REGION Network 107: DB34.DBB10 -> DB86.DBB20 / 8 y 8
   // Falla Compresor ABC2 Baja Presion de Agua
   // Falla Compresor ABC2 Alta Temperatura de Aire
   // Falla Compresor ABC2 Alta Temperatura de agua
   // Falla Compresor ABC3 Baja Presion de Aceite
   // Falla Compresor ABC3 Baja Presion de Agua
   // Falla Compresor ABC3 Alta Temperatura de Aire
   // Falla Compresor ABC3 Alta Temperatura de agua
   // Falla Compresor ABC4 Baja Presion de Aceite
   RUNG wire#powerrail
      { S7_GenerateENO := "TRUE" } Move(in := %DB34.DBB10, out1 => %DB86.DBB20)
      "And-Byte MTA"(IN0 := %DB86.DBB21, IN1 := %DB34.DBB10, OUT2 => %DB86.DBB21)
      { S7_GenerateENO := "TRUE" } Move(in := %DB86.DBB21, out1 => %DB35.DBB10)
   END_RUNG
   // the same network as SCL:
   // ENO of a box is taken as its EN; it also drops when the box reports an error
   %DB86.DBB20 := %DB34.DBB10;
   "And-Byte MTA"(IN0 := %DB86.DBB21, IN1 := %DB34.DBB10, OUT2 => %DB86.DBB21, ENO => #_w1);
   IF #_w1 THEN %DB35.DBB10 := %DB86.DBB21; END_IF;
END_REGION

REGION Network 108: DB34.DBB11 -> DB86.DBB22 / 8 y 8
   // Falla Compresor ABC4 Alta Temperatura de Aire
   // Falla Compresor ABC4 Alta Temperatura de Aire
   // Falla Compresor ABC4 Alta Temperatura de agua
   // Falla Compresor ABC5 Baja Presion de Aceite
   // Falla Compresor ABC5 Alta Temperatura de Aire
   // Falla Compresor ABC5 Alta Temperatura de Aire
   // Falla Compresor ABC5 Alta Temperatura de agua
   // Falla Compresor Bellis & MHW28 Baja Presion Aceite
   RUNG wire#powerrail
      { S7_GenerateENO := "TRUE" } Move(in := %DB34.DBB11, out1 => %DB86.DBB22)
      "And-Byte MTA"(IN0 := %DB86.DBB23, IN1 := %DB34.DBB11, OUT2 => %DB86.DBB23)
      { S7_GenerateENO := "TRUE" } Move(in := %DB86.DBB23, out1 => %DB35.DBB11)
   END_RUNG
   // the same network as SCL:
   // ENO of a box is taken as its EN; it also drops when the box reports an error
   %DB86.DBB22 := %DB34.DBB11;
   "And-Byte MTA"(IN0 := %DB86.DBB23, IN1 := %DB34.DBB11, OUT2 => %DB86.DBB23, ENO => #_w1);
   IF #_w1 THEN %DB35.DBB11 := %DB86.DBB23; END_IF;
END_REGION

REGION Network 109: DB34.DBB12 -> DB86.DBB24 / 8 y 8
   // Falla Compresor Bellis & MHW28 Baja Presion de Agua
   // Falla Compresor Bellis & MHW28 Alta temperatura de Aire
   // Falla Compresor Bellis & MHW28 Alta temperatura de Agua
   // Falla Compresor Bellis & MHW28 Falla de Flujostato
   // Requiere Marcha MC001
   // Requiere Marcha MC002
   // Requiere Marcha MC003
   // Requiere Marcha MC004
   RUNG wire#powerrail
      { S7_GenerateENO := "TRUE" } Move(in := %DB34.DBB12, out1 => %DB86.DBB24)
      "And-Byte MTA"(IN0 := %DB86.DBB25, IN1 := %DB34.DBB12, OUT2 => %DB86.DBB25)
      { S7_GenerateENO := "TRUE" } Move(in := %DB86.DBB25, out1 => %DB35.DBB12)
   END_RUNG
   // the same network as SCL:
   // ENO of a box is taken as its EN; it also drops when the box reports an error
   %DB86.DBB24 := %DB34.DBB12;
   "And-Byte MTA"(IN0 := %DB86.DBB25, IN1 := %DB34.DBB12, OUT2 => %DB86.DBB25, ENO => #_w1);
   IF #_w1 THEN %DB35.DBB12 := %DB86.DBB25; END_IF;
END_REGION

REGION Network 110: DB34.DBB13 -> DB86.DBB26 / 8 y 8
   // Requiere Marcha MC005
   // Falla Conexión con sensor de Temperatura torres de Cavaleto
   // Falla Conexión con sensor de Temperatura torres de Chillers
   // Falla Conexión con sensor de Presión de ALTA
   // Falla Conexión con sensor de Presión de ALTA redundante
   // Falla Conexión con sensor de Presión de Baja
   // Falla Presión de Alta en Límite Mínimo
   // Falla Presión de Alta en demasiado Baja
   RUNG wire#powerrail
      { S7_GenerateENO := "TRUE" } Move(in := %DB34.DBB13, out1 => %DB86.DBB26)
      "And-Byte MTA"(IN0 := %DB86.DBB27, IN1 := %DB34.DBB13, OUT2 => %DB86.DBB27)
      { S7_GenerateENO := "TRUE" } Move(in := %DB86.DBB27, out1 => %DB35.DBB13)
   END_RUNG
   // the same network as SCL:
   // ENO of a box is taken as its EN; it also drops when the box reports an error
   %DB86.DBB26 := %DB34.DBB13;
   "And-Byte MTA"(IN0 := %DB86.DBB27, IN1 := %DB34.DBB13, OUT2 => %DB86.DBB27, ENO => #_w1);
   IF #_w1 THEN %DB35.DBB13 := %DB86.DBB27; END_IF;
END_REGION

REGION Network 111: DB34.DBB14 -> DB86.DBB28 / 8 y 8
   // Falla Presión de Alta en demasiado Alta
   // Falla Presión de Alta en Límite Máximo
   // Falla Presión de Baja en Límite Mínimo
   // Falla Presión de Baja en demasiado Baja
   // Falla Presión de Baja en demasiado Alta
   // Falla Presión de Baja en Límite Máximo
   // Falla en chiller de envasado chico
   // Falla en chiller de soplado chico
   RUNG wire#powerrail
      { S7_GenerateENO := "TRUE" } Move(in := %DB34.DBB14, out1 => %DB86.DBB28)
      "And-Byte MTA"(IN0 := %DB86.DBB29, IN1 := %DB34.DBB14, OUT2 => %DB86.DBB29)
      { S7_GenerateENO := "TRUE" } Move(in := %DB86.DBB29, out1 => %DB35.DBB14)
   END_RUNG
   // the same network as SCL:
   // ENO of a box is taken as its EN; it also drops when the box reports an error
   %DB86.DBB28 := %DB34.DBB14;
   "And-Byte MTA"(IN0 := %DB86.DBB29, IN1 := %DB34.DBB14, OUT2 => %DB86.DBB29, ENO => #_w1);
   IF #_w1 THEN %DB35.DBB14 := %DB86.DBB29; END_IF;
END_REGION

REGION Network 112: DB34.DBB15 -> DB86.DBB30 / 8 y 8
   // Horas máximas en Compresor 1
   // Horas máximas en Compresor 2
   // Horas máximas en Compresor 3
   // Horas máximas en Compresor 4
   // Horas máximas en Compresor 5
   // Falla algún contactor en Booster 1
   // Falla algún guardamotor en Booster 1
   // Presión Alta en Booster
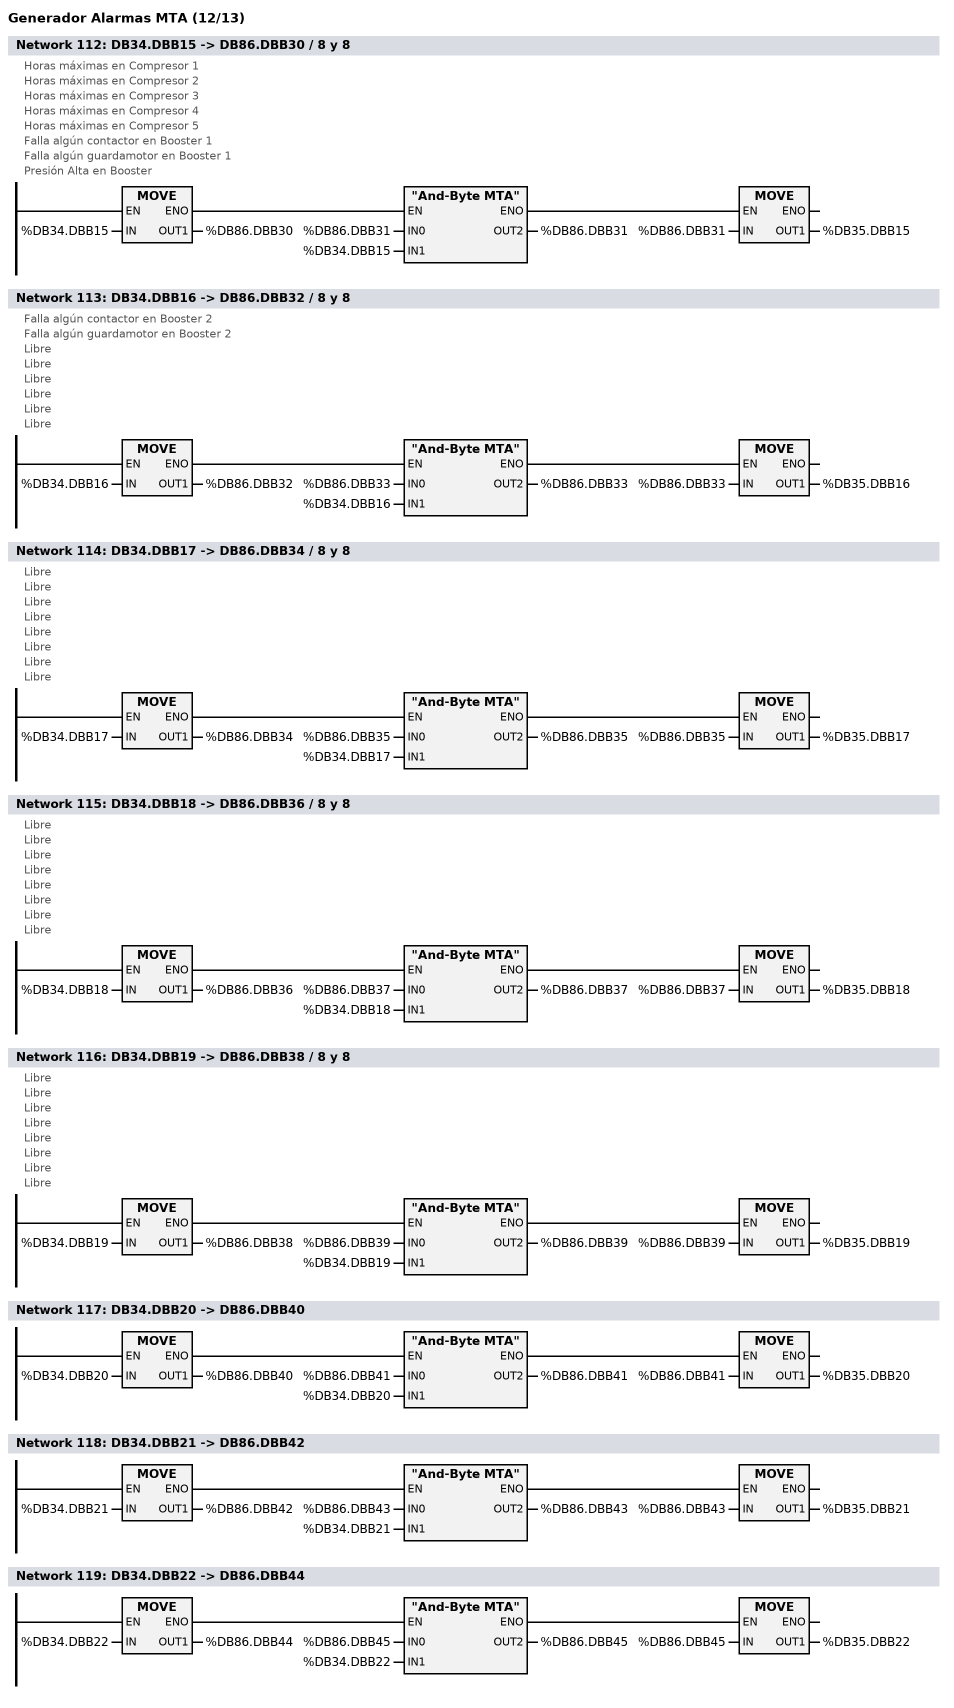
   RUNG wire#powerrail
      { S7_GenerateENO := "TRUE" } Move(in := %DB34.DBB15, out1 => %DB86.DBB30)
      "And-Byte MTA"(IN0 := %DB86.DBB31, IN1 := %DB34.DBB15, OUT2 => %DB86.DBB31)
      { S7_GenerateENO := "TRUE" } Move(in := %DB86.DBB31, out1 => %DB35.DBB15)
   END_RUNG
   // the same network as SCL:
   // ENO of a box is taken as its EN; it also drops when the box reports an error
   %DB86.DBB30 := %DB34.DBB15;
   "And-Byte MTA"(IN0 := %DB86.DBB31, IN1 := %DB34.DBB15, OUT2 => %DB86.DBB31, ENO => #_w1);
   IF #_w1 THEN %DB35.DBB15 := %DB86.DBB31; END_IF;
END_REGION

REGION Network 113: DB34.DBB16 -> DB86.DBB32 / 8 y 8
   // Falla algún contactor en Booster 2
   // Falla algún guardamotor en Booster 2
   // Libre
   // Libre
   // Libre
   // Libre
   // Libre
   // Libre
   RUNG wire#powerrail
      { S7_GenerateENO := "TRUE" } Move(in := %DB34.DBB16, out1 => %DB86.DBB32)
      "And-Byte MTA"(IN0 := %DB86.DBB33, IN1 := %DB34.DBB16, OUT2 => %DB86.DBB33)
      { S7_GenerateENO := "TRUE" } Move(in := %DB86.DBB33, out1 => %DB35.DBB16)
   END_RUNG
   // the same network as SCL:
   // ENO of a box is taken as its EN; it also drops when the box reports an error
   %DB86.DBB32 := %DB34.DBB16;
   "And-Byte MTA"(IN0 := %DB86.DBB33, IN1 := %DB34.DBB16, OUT2 => %DB86.DBB33, ENO => #_w1);
   IF #_w1 THEN %DB35.DBB16 := %DB86.DBB33; END_IF;
END_REGION

REGION Network 114: DB34.DBB17 -> DB86.DBB34 / 8 y 8
   // Libre
   // Libre
   // Libre
   // Libre
   // Libre
   // Libre
   // Libre
   // Libre
   RUNG wire#powerrail
      { S7_GenerateENO := "TRUE" } Move(in := %DB34.DBB17, out1 => %DB86.DBB34)
      "And-Byte MTA"(IN0 := %DB86.DBB35, IN1 := %DB34.DBB17, OUT2 => %DB86.DBB35)
      { S7_GenerateENO := "TRUE" } Move(in := %DB86.DBB35, out1 => %DB35.DBB17)
   END_RUNG
   // the same network as SCL:
   // ENO of a box is taken as its EN; it also drops when the box reports an error
   %DB86.DBB34 := %DB34.DBB17;
   "And-Byte MTA"(IN0 := %DB86.DBB35, IN1 := %DB34.DBB17, OUT2 => %DB86.DBB35, ENO => #_w1);
   IF #_w1 THEN %DB35.DBB17 := %DB86.DBB35; END_IF;
END_REGION

REGION Network 115: DB34.DBB18 -> DB86.DBB36 / 8 y 8
   // Libre
   // Libre
   // Libre
   // Libre
   // Libre
   // Libre
   // Libre
   // Libre
   RUNG wire#powerrail
      { S7_GenerateENO := "TRUE" } Move(in := %DB34.DBB18, out1 => %DB86.DBB36)
      "And-Byte MTA"(IN0 := %DB86.DBB37, IN1 := %DB34.DBB18, OUT2 => %DB86.DBB37)
      { S7_GenerateENO := "TRUE" } Move(in := %DB86.DBB37, out1 => %DB35.DBB18)
   END_RUNG
   // the same network as SCL:
   // ENO of a box is taken as its EN; it also drops when the box reports an error
   %DB86.DBB36 := %DB34.DBB18;
   "And-Byte MTA"(IN0 := %DB86.DBB37, IN1 := %DB34.DBB18, OUT2 => %DB86.DBB37, ENO => #_w1);
   IF #_w1 THEN %DB35.DBB18 := %DB86.DBB37; END_IF;
END_REGION

REGION Network 116: DB34.DBB19 -> DB86.DBB38 / 8 y 8
   // Libre
   // Libre
   // Libre
   // Libre
   // Libre
   // Libre
   // Libre
   // Libre
   RUNG wire#powerrail
      { S7_GenerateENO := "TRUE" } Move(in := %DB34.DBB19, out1 => %DB86.DBB38)
      "And-Byte MTA"(IN0 := %DB86.DBB39, IN1 := %DB34.DBB19, OUT2 => %DB86.DBB39)
      { S7_GenerateENO := "TRUE" } Move(in := %DB86.DBB39, out1 => %DB35.DBB19)
   END_RUNG
   // the same network as SCL:
   // ENO of a box is taken as its EN; it also drops when the box reports an error
   %DB86.DBB38 := %DB34.DBB19;
   "And-Byte MTA"(IN0 := %DB86.DBB39, IN1 := %DB34.DBB19, OUT2 => %DB86.DBB39, ENO => #_w1);
   IF #_w1 THEN %DB35.DBB19 := %DB86.DBB39; END_IF;
END_REGION

REGION Network 117: DB34.DBB20 -> DB86.DBB40
   RUNG wire#powerrail
      { S7_GenerateENO := "TRUE" } Move(in := %DB34.DBB20, out1 => %DB86.DBB40)
      "And-Byte MTA"(IN0 := %DB86.DBB41, IN1 := %DB34.DBB20, OUT2 => %DB86.DBB41)
      { S7_GenerateENO := "TRUE" } Move(in := %DB86.DBB41, out1 => %DB35.DBB20)
   END_RUNG
   // the same network as SCL:
   // ENO of a box is taken as its EN; it also drops when the box reports an error
   %DB86.DBB40 := %DB34.DBB20;
   "And-Byte MTA"(IN0 := %DB86.DBB41, IN1 := %DB34.DBB20, OUT2 => %DB86.DBB41, ENO => #_w1);
   IF #_w1 THEN %DB35.DBB20 := %DB86.DBB41; END_IF;
END_REGION

REGION Network 118: DB34.DBB21 -> DB86.DBB42
   RUNG wire#powerrail
      { S7_GenerateENO := "TRUE" } Move(in := %DB34.DBB21, out1 => %DB86.DBB42)
      "And-Byte MTA"(IN0 := %DB86.DBB43, IN1 := %DB34.DBB21, OUT2 => %DB86.DBB43)
      { S7_GenerateENO := "TRUE" } Move(in := %DB86.DBB43, out1 => %DB35.DBB21)
   END_RUNG
   // the same network as SCL:
   // ENO of a box is taken as its EN; it also drops when the box reports an error
   %DB86.DBB42 := %DB34.DBB21;
   "And-Byte MTA"(IN0 := %DB86.DBB43, IN1 := %DB34.DBB21, OUT2 => %DB86.DBB43, ENO => #_w1);
   IF #_w1 THEN %DB35.DBB21 := %DB86.DBB43; END_IF;
END_REGION

REGION Network 119: DB34.DBB22 -> DB86.DBB44
   RUNG wire#powerrail
      { S7_GenerateENO := "TRUE" } Move(in := %DB34.DBB22, out1 => %DB86.DBB44)
      "And-Byte MTA"(IN0 := %DB86.DBB45, IN1 := %DB34.DBB22, OUT2 => %DB86.DBB45)
      { S7_GenerateENO := "TRUE" } Move(in := %DB86.DBB45, out1 => %DB35.DBB22)
   END_RUNG
   // the same network as SCL:
   // ENO of a box is taken as its EN; it also drops when the box reports an error
   %DB86.DBB44 := %DB34.DBB22;
   "And-Byte MTA"(IN0 := %DB86.DBB45, IN1 := %DB34.DBB22, OUT2 => %DB86.DBB45, ENO => #_w1);
   IF #_w1 THEN %DB35.DBB22 := %DB86.DBB45; END_IF;
END_REGION

REGION Network 120: DB34.DBB23 -> DB86.DBB46
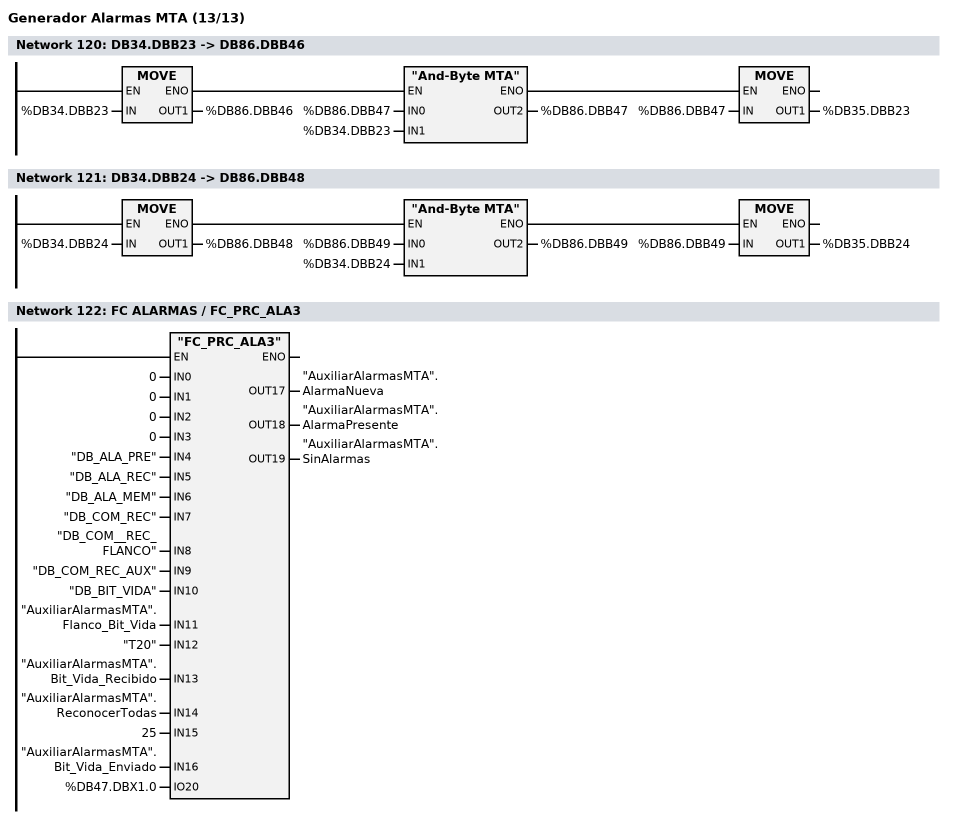
   RUNG wire#powerrail
      { S7_GenerateENO := "TRUE" } Move(in := %DB34.DBB23, out1 => %DB86.DBB46)
      "And-Byte MTA"(IN0 := %DB86.DBB47, IN1 := %DB34.DBB23, OUT2 => %DB86.DBB47)
      { S7_GenerateENO := "TRUE" } Move(in := %DB86.DBB47, out1 => %DB35.DBB23)
   END_RUNG
   // the same network as SCL:
   // ENO of a box is taken as its EN; it also drops when the box reports an error
   %DB86.DBB46 := %DB34.DBB23;
   "And-Byte MTA"(IN0 := %DB86.DBB47, IN1 := %DB34.DBB23, OUT2 => %DB86.DBB47, ENO => #_w1);
   IF #_w1 THEN %DB35.DBB23 := %DB86.DBB47; END_IF;
END_REGION

REGION Network 121: DB34.DBB24 -> DB86.DBB48
   RUNG wire#powerrail
      { S7_GenerateENO := "TRUE" } Move(in := %DB34.DBB24, out1 => %DB86.DBB48)
      "And-Byte MTA"(IN0 := %DB86.DBB49, IN1 := %DB34.DBB24, OUT2 => %DB86.DBB49)
      { S7_GenerateENO := "TRUE" } Move(in := %DB86.DBB49, out1 => %DB35.DBB24)
   END_RUNG
   // the same network as SCL:
   // ENO of a box is taken as its EN; it also drops when the box reports an error
   %DB86.DBB48 := %DB34.DBB24;
   "And-Byte MTA"(IN0 := %DB86.DBB49, IN1 := %DB34.DBB24, OUT2 => %DB86.DBB49, ENO => #_w1);
   IF #_w1 THEN %DB35.DBB24 := %DB86.DBB49; END_IF;
END_REGION

REGION Network 122: FC ALARMAS / FC_PRC_ALA3
   RUNG wire#powerrail
      "FC_PRC_ALA3"(IN0 := 0, IN1 := 0, IN2 := 0, IN3 := 0, IN4 := "DB_ALA_PRE", IN5 := "DB_ALA_REC", IN6 := "DB_ALA_MEM", IN7 := "DB_COM_REC", IN8 := "DB_COM__REC_FLANCO", IN9 := "DB_COM_REC_AUX", IN10 := "DB_BIT_VIDA", IN11 := "AuxiliarAlarmasMTA".Flanco_Bit_Vida, IN12 := "T20", IN13 := "AuxiliarAlarmasMTA".Bit_Vida_Recibido, IN14 := "AuxiliarAlarmasMTA".ReconocerTodas, IN15 := 25, IN16 := "AuxiliarAlarmasMTA".Bit_Vida_Enviado, IO20 := %DB47.DBX1.0, OUT17 => "AuxiliarAlarmasMTA".AlarmaNueva, OUT18 => "AuxiliarAlarmasMTA".AlarmaPresente, OUT19 => "AuxiliarAlarmasMTA".SinAlarmas)
   END_RUNG
   // the same network as SCL:
   "FC_PRC_ALA3"(IN0 := 0,
                 IN1 := 0,
                 IN2 := 0,
                 IN3 := 0,
                 IN4 := "DB_ALA_PRE",
                 IN5 := "DB_ALA_REC",
                 IN6 := "DB_ALA_MEM",
                 IN7 := "DB_COM_REC",
                 IN8 := "DB_COM__REC_FLANCO",
                 IN9 := "DB_COM_REC_AUX",
                 IN10 := "DB_BIT_VIDA",
                 IN11 := "AuxiliarAlarmasMTA".Flanco_Bit_Vida,
                 IN12 := "T20",
                 IN13 := "AuxiliarAlarmasMTA".Bit_Vida_Recibido,
                 IN14 := "AuxiliarAlarmasMTA".ReconocerTodas,
                 IN15 := 25,
                 IN16 := "AuxiliarAlarmasMTA".Bit_Vida_Enviado,
                 IO20 := %DB47.DBX1.0,
                 OUT17 => "AuxiliarAlarmasMTA".AlarmaNueva,
                 OUT18 => "AuxiliarAlarmasMTA".AlarmaPresente,
                 OUT19 => "AuxiliarAlarmasMTA".SinAlarmas);
END_REGION
END_FUNCTION

FUNCTION "FalCmpAlta" : Void   // FC49, LAD
{ S7_Optimized_Access := 'FALSE' }
VERSION : 0.1
   VAR_TEMP   // added for the SCL form of the ladder/FBD networks
      _w1 : Bool;
      _w2 : Bool;
      _s5time1 : S5Time;
   END_VAR
BEGIN

REGION Network 1: Fallas de MC001 - Compresor de Alta ABC2
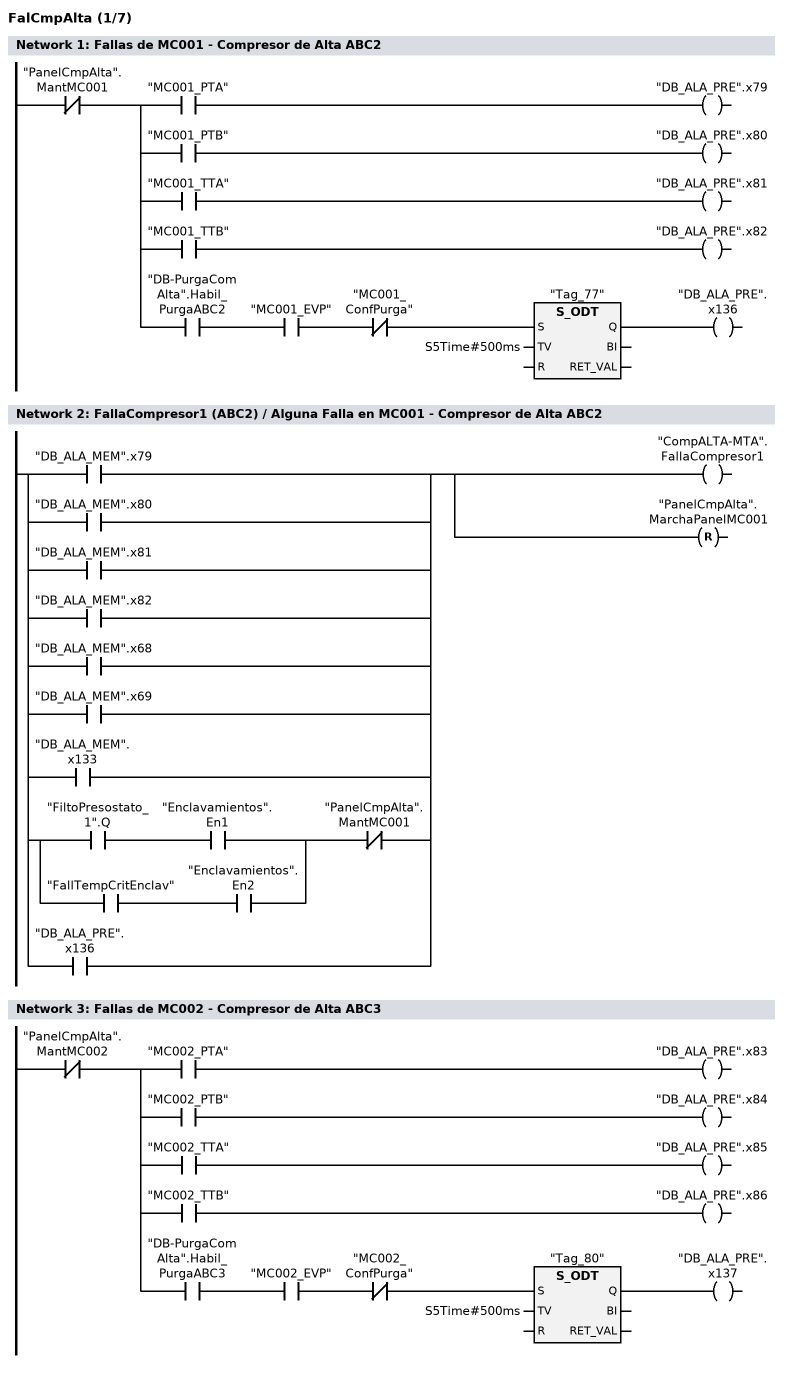
   RUNG wire#powerrail
      I_Contact( "PanelCmpAlta".MantMC001 )
      wire#w1
      Contact( "MC001_PTA" )
      Coil( "DB_ALA_PRE".x79 )
   END_RUNG
   RUNG wire#w1
      Contact( "MC001_PTB" )
      Coil( "DB_ALA_PRE".x80 )
   END_RUNG
   RUNG wire#w1
      Contact( "MC001_TTA" )
      Coil( "DB_ALA_PRE".x81 )
   END_RUNG
   RUNG wire#w1
      Contact( "MC001_TTB" )
      Coil( "DB_ALA_PRE".x82 )
   END_RUNG
   RUNG wire#w1
      Contact( "DB-PurgaComAlta".Habil_PurgaABC2 )
      Contact( "MC001_EVP" )
      I_Contact( "MC001_ConfPurga" )
      S_ODT(T_NO := "Tag_77", TV := S5Time#500ms, R :=, BI =>, RET_VAL =>)
      Coil( "DB_ALA_PRE".x136 )
   END_RUNG
   // the same network as SCL:
   #_w1 := NOT "PanelCmpAlta".MantMC001;
   "DB_ALA_PRE".x79 := #_w1 AND "MC001_PTA";
   "DB_ALA_PRE".x80 := #_w1 AND "MC001_PTB";
   "DB_ALA_PRE".x81 := #_w1 AND "MC001_TTA";
   "DB_ALA_PRE".x82 := #_w1 AND "MC001_TTB";
   #_s5time1 := S_ODT(T_NO := "Tag_77",
                      S := #_w1 AND "DB-PurgaComAlta".Habil_PurgaABC2 AND "MC001_EVP" AND NOT "MC001_ConfPurga",
                      TV := S5Time#500ms,
                      Q => #_w2);
   "DB_ALA_PRE".x136 := #_w2;
END_REGION

REGION Network 2: FallaCompresor1 (ABC2) / Alguna Falla en MC001 - Compresor de Alta ABC2
   RUNG wire#powerrail
      Contact( "DB_ALA_MEM".x79 )
      wire#w1
      Coil( "CompALTA-MTA".FallaCompresor1 )
   END_RUNG
   RUNG wire#powerrail
      Contact( "DB_ALA_MEM".x80 )
   END_RUNG wire#w1
   RUNG wire#powerrail
      Contact( "DB_ALA_MEM".x81 )
   END_RUNG wire#w1
   RUNG wire#powerrail
      Contact( "DB_ALA_MEM".x82 )
   END_RUNG wire#w1
   RUNG wire#powerrail
      Contact( "DB_ALA_MEM".x68 )
   END_RUNG wire#w1
   RUNG wire#powerrail
      Contact( "DB_ALA_MEM".x69 )
   END_RUNG wire#w1
   RUNG wire#powerrail
      Contact( "DB_ALA_MEM".x133 )
   END_RUNG wire#w1
   RUNG wire#powerrail
      Contact( "FiltoPresostato_1".Q )
      Contact( "Enclavamientos".En1 )
      wire#w2
      I_Contact( "PanelCmpAlta".MantMC001 )
   END_RUNG wire#w1
   RUNG wire#powerrail
      Contact( "FallTempCritEnclav" )
      Contact( "Enclavamientos".En2 )
   END_RUNG wire#w2
   RUNG wire#powerrail
      Contact( "DB_ALA_PRE".x136 )
   END_RUNG wire#w1
   RUNG wire#w1
      R_Coil( "PanelCmpAlta".MarchaPanelMC001 )
   END_RUNG
   // the same network as SCL:
   "CompALTA-MTA".FallaCompresor1 := "DB_ALA_MEM".x79 OR "DB_ALA_MEM".x80 OR "DB_ALA_MEM".x81 OR "DB_ALA_MEM".x82 OR "DB_ALA_MEM".x68 OR "DB_ALA_MEM".x69 OR "DB_ALA_MEM".x133 OR ((("FiltoPresostato_1".Q AND "Enclavamientos".En1) OR ("FallTempCritEnclav" AND "Enclavamientos".En2)) AND NOT "PanelCmpAlta".MantMC001) OR "DB_ALA_PRE".x136;
   IF "CompALTA-MTA".FallaCompresor1 THEN "PanelCmpAlta".MarchaPanelMC001 := FALSE; END_IF;
END_REGION

REGION Network 3: Fallas de MC002 - Compresor de Alta ABC3
   RUNG wire#powerrail
      I_Contact( "PanelCmpAlta".MantMC002 )
      wire#w1
      Contact( "MC002_PTA" )
      Coil( "DB_ALA_PRE".x83 )
   END_RUNG
   RUNG wire#w1
      Contact( "MC002_PTB" )
      Coil( "DB_ALA_PRE".x84 )
   END_RUNG
   RUNG wire#w1
      Contact( "MC002_TTA" )
      Coil( "DB_ALA_PRE".x85 )
   END_RUNG
   RUNG wire#w1
      Contact( "MC002_TTB" )
      Coil( "DB_ALA_PRE".x86 )
   END_RUNG
   RUNG wire#w1
      Contact( "DB-PurgaComAlta".Habil_PurgaABC3 )
      Contact( "MC002_EVP" )
      I_Contact( "MC002_ConfPurga" )
      S_ODT(T_NO := "Tag_80", TV := S5Time#500ms, R :=, BI =>, RET_VAL =>)
      Coil( "DB_ALA_PRE".x137 )
   END_RUNG
   // the same network as SCL:
   #_w1 := NOT "PanelCmpAlta".MantMC002;
   "DB_ALA_PRE".x83 := #_w1 AND "MC002_PTA";
   "DB_ALA_PRE".x84 := #_w1 AND "MC002_PTB";
   "DB_ALA_PRE".x85 := #_w1 AND "MC002_TTA";
   "DB_ALA_PRE".x86 := #_w1 AND "MC002_TTB";
   #_s5time1 := S_ODT(T_NO := "Tag_80",
                      S := #_w1 AND "DB-PurgaComAlta".Habil_PurgaABC3 AND "MC002_EVP" AND NOT "MC002_ConfPurga",
                      TV := S5Time#500ms,
                      Q => #_w2);
   "DB_ALA_PRE".x137 := #_w2;
END_REGION

REGION Network 4: FallaCompresor2 (ABC3) / Alguna Falla en MC002 - Compresor de Alta ABC3
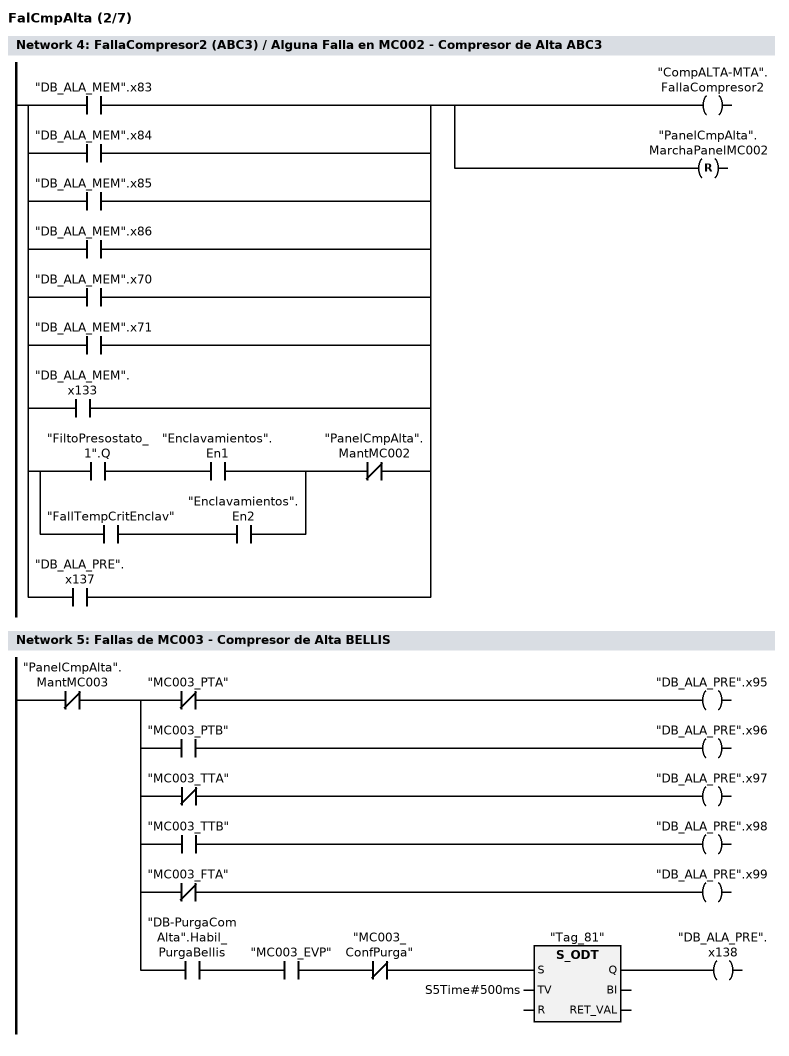
   RUNG wire#powerrail
      Contact( "DB_ALA_MEM".x83 )
      wire#w1
      Coil( "CompALTA-MTA".FallaCompresor2 )
   END_RUNG
   RUNG wire#powerrail
      Contact( "DB_ALA_MEM".x84 )
   END_RUNG wire#w1
   RUNG wire#powerrail
      Contact( "DB_ALA_MEM".x85 )
   END_RUNG wire#w1
   RUNG wire#powerrail
      Contact( "DB_ALA_MEM".x86 )
   END_RUNG wire#w1
   RUNG wire#powerrail
      Contact( "DB_ALA_MEM".x70 )
   END_RUNG wire#w1
   RUNG wire#powerrail
      Contact( "DB_ALA_MEM".x71 )
   END_RUNG wire#w1
   RUNG wire#powerrail
      Contact( "DB_ALA_MEM".x133 )
   END_RUNG wire#w1
   RUNG wire#powerrail
      Contact( "FiltoPresostato_1".Q )
      Contact( "Enclavamientos".En1 )
      wire#w2
      I_Contact( "PanelCmpAlta".MantMC002 )
   END_RUNG wire#w1
   RUNG wire#powerrail
      Contact( "FallTempCritEnclav" )
      Contact( "Enclavamientos".En2 )
   END_RUNG wire#w2
   RUNG wire#powerrail
      Contact( "DB_ALA_PRE".x137 )
   END_RUNG wire#w1
   RUNG wire#w1
      R_Coil( "PanelCmpAlta".MarchaPanelMC002 )
   END_RUNG
   // the same network as SCL:
   "CompALTA-MTA".FallaCompresor2 := "DB_ALA_MEM".x83 OR "DB_ALA_MEM".x84 OR "DB_ALA_MEM".x85 OR "DB_ALA_MEM".x86 OR "DB_ALA_MEM".x70 OR "DB_ALA_MEM".x71 OR "DB_ALA_MEM".x133 OR ((("FiltoPresostato_1".Q AND "Enclavamientos".En1) OR ("FallTempCritEnclav" AND "Enclavamientos".En2)) AND NOT "PanelCmpAlta".MantMC002) OR "DB_ALA_PRE".x137;
   IF "CompALTA-MTA".FallaCompresor2 THEN "PanelCmpAlta".MarchaPanelMC002 := FALSE; END_IF;
END_REGION

REGION Network 5: Fallas de MC003 - Compresor de Alta BELLIS
   RUNG wire#powerrail
      I_Contact( "PanelCmpAlta".MantMC003 )
      wire#w1
      I_Contact( "MC003_PTA" )
      Coil( "DB_ALA_PRE".x95 )
   END_RUNG
   RUNG wire#w1
      Contact( "MC003_PTB" )
      Coil( "DB_ALA_PRE".x96 )
   END_RUNG
   RUNG wire#w1
      I_Contact( "MC003_TTA" )
      Coil( "DB_ALA_PRE".x97 )
   END_RUNG
   RUNG wire#w1
      Contact( "MC003_TTB" )
      Coil( "DB_ALA_PRE".x98 )
   END_RUNG
   RUNG wire#w1
      I_Contact( "MC003_FTA" )
      Coil( "DB_ALA_PRE".x99 )
   END_RUNG
   RUNG wire#w1
      Contact( "DB-PurgaComAlta".Habil_PurgaBellis )
      Contact( "MC003_EVP" )
      I_Contact( "MC003_ConfPurga" )
      S_ODT(T_NO := "Tag_81", TV := S5Time#500ms, R :=, BI =>, RET_VAL =>)
      Coil( "DB_ALA_PRE".x138 )
   END_RUNG
   // the same network as SCL:
   #_w1 := NOT "PanelCmpAlta".MantMC003;
   "DB_ALA_PRE".x95 := #_w1 AND NOT "MC003_PTA";
   "DB_ALA_PRE".x96 := #_w1 AND "MC003_PTB";
   "DB_ALA_PRE".x97 := #_w1 AND NOT "MC003_TTA";
   "DB_ALA_PRE".x98 := #_w1 AND "MC003_TTB";
   "DB_ALA_PRE".x99 := #_w1 AND NOT "MC003_FTA";
   #_s5time1 := S_ODT(T_NO := "Tag_81",
                      S := #_w1 AND "DB-PurgaComAlta".Habil_PurgaBellis AND "MC003_EVP" AND NOT "MC003_ConfPurga",
                      TV := S5Time#500ms,
                      Q => #_w2);
   "DB_ALA_PRE".x138 := #_w2;
END_REGION

REGION Network 6: FallaCompresor3 (Bellis) / Alguna Falla en MC003 - Compresor de Alta BELLIS
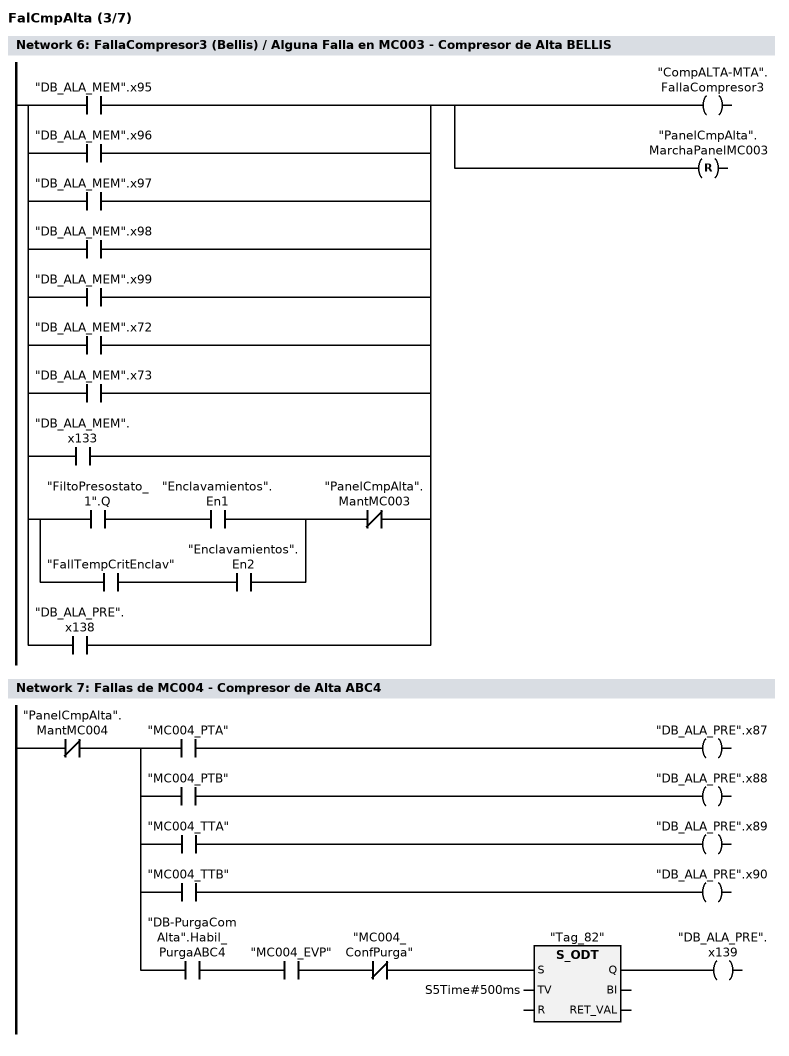
   RUNG wire#powerrail
      Contact( "DB_ALA_MEM".x95 )
      wire#w1
      Coil( "CompALTA-MTA".FallaCompresor3 )
   END_RUNG
   RUNG wire#powerrail
      Contact( "DB_ALA_MEM".x96 )
   END_RUNG wire#w1
   RUNG wire#powerrail
      Contact( "DB_ALA_MEM".x97 )
   END_RUNG wire#w1
   RUNG wire#powerrail
      Contact( "DB_ALA_MEM".x98 )
   END_RUNG wire#w1
   RUNG wire#powerrail
      Contact( "DB_ALA_MEM".x99 )
   END_RUNG wire#w1
   RUNG wire#powerrail
      Contact( "DB_ALA_MEM".x72 )
   END_RUNG wire#w1
   RUNG wire#powerrail
      Contact( "DB_ALA_MEM".x73 )
   END_RUNG wire#w1
   RUNG wire#powerrail
      Contact( "DB_ALA_MEM".x133 )
   END_RUNG wire#w1
   RUNG wire#powerrail
      Contact( "FiltoPresostato_1".Q )
      Contact( "Enclavamientos".En1 )
      wire#w2
      I_Contact( "PanelCmpAlta".MantMC003 )
   END_RUNG wire#w1
   RUNG wire#powerrail
      Contact( "FallTempCritEnclav" )
      Contact( "Enclavamientos".En2 )
   END_RUNG wire#w2
   RUNG wire#powerrail
      Contact( "DB_ALA_PRE".x138 )
   END_RUNG wire#w1
   RUNG wire#w1
      R_Coil( "PanelCmpAlta".MarchaPanelMC003 )
   END_RUNG
   // the same network as SCL:
   "CompALTA-MTA".FallaCompresor3 := "DB_ALA_MEM".x95 OR "DB_ALA_MEM".x96 OR "DB_ALA_MEM".x97 OR "DB_ALA_MEM".x98 OR "DB_ALA_MEM".x99 OR "DB_ALA_MEM".x72 OR "DB_ALA_MEM".x73 OR "DB_ALA_MEM".x133 OR ((("FiltoPresostato_1".Q AND "Enclavamientos".En1) OR ("FallTempCritEnclav" AND "Enclavamientos".En2)) AND NOT "PanelCmpAlta".MantMC003) OR "DB_ALA_PRE".x138;
   IF "CompALTA-MTA".FallaCompresor3 THEN "PanelCmpAlta".MarchaPanelMC003 := FALSE; END_IF;
END_REGION

REGION Network 7: Fallas de MC004 - Compresor de Alta ABC4
   RUNG wire#powerrail
      I_Contact( "PanelCmpAlta".MantMC004 )
      wire#w1
      Contact( "MC004_PTA" )
      Coil( "DB_ALA_PRE".x87 )
   END_RUNG
   RUNG wire#w1
      Contact( "MC004_PTB" )
      Coil( "DB_ALA_PRE".x88 )
   END_RUNG
   RUNG wire#w1
      Contact( "MC004_TTA" )
      Coil( "DB_ALA_PRE".x89 )
   END_RUNG
   RUNG wire#w1
      Contact( "MC004_TTB" )
      Coil( "DB_ALA_PRE".x90 )
   END_RUNG
   RUNG wire#w1
      Contact( "DB-PurgaComAlta".Habil_PurgaABC4 )
      Contact( "MC004_EVP" )
      I_Contact( "MC004_ConfPurga" )
      S_ODT(T_NO := "Tag_82", TV := S5Time#500ms, R :=, BI =>, RET_VAL =>)
      Coil( "DB_ALA_PRE".x139 )
   END_RUNG
   // the same network as SCL:
   #_w1 := NOT "PanelCmpAlta".MantMC004;
   "DB_ALA_PRE".x87 := #_w1 AND "MC004_PTA";
   "DB_ALA_PRE".x88 := #_w1 AND "MC004_PTB";
   "DB_ALA_PRE".x89 := #_w1 AND "MC004_TTA";
   "DB_ALA_PRE".x90 := #_w1 AND "MC004_TTB";
   #_s5time1 := S_ODT(T_NO := "Tag_82",
                      S := #_w1 AND "DB-PurgaComAlta".Habil_PurgaABC4 AND "MC004_EVP" AND NOT "MC004_ConfPurga",
                      TV := S5Time#500ms,
                      Q => #_w2);
   "DB_ALA_PRE".x139 := #_w2;
END_REGION

REGION Network 8: FallaCompresor4 (ABC4) / Alguna Falla en MC004 - Compresor de Alta ABC4
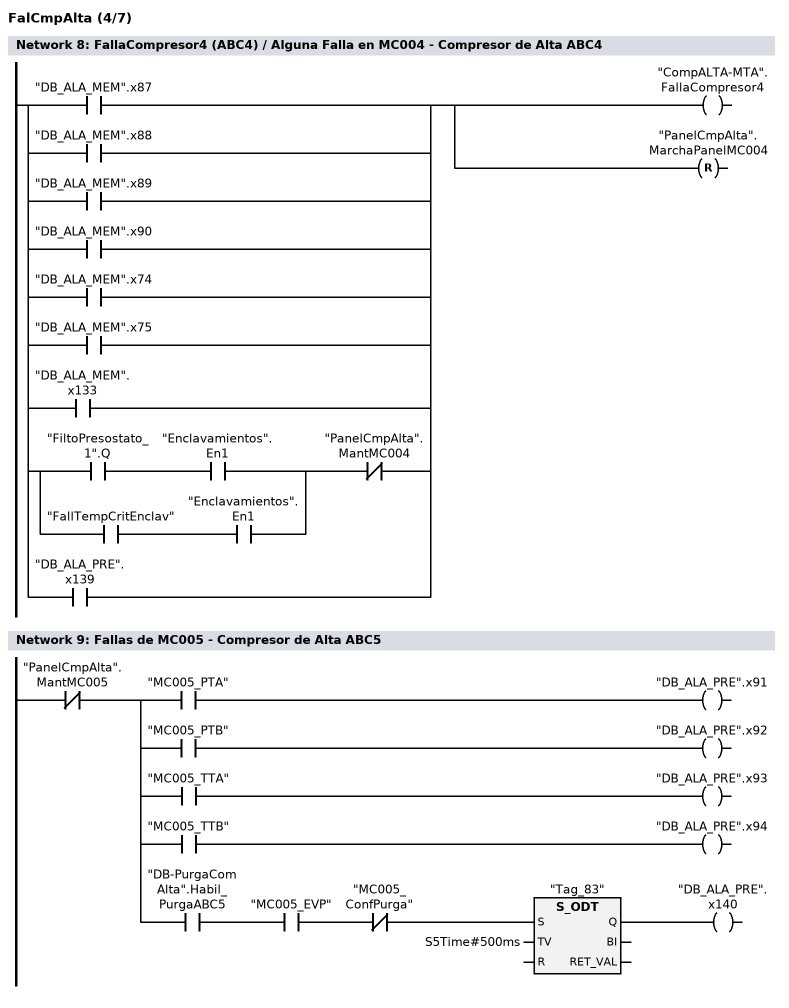
   RUNG wire#powerrail
      Contact( "DB_ALA_MEM".x87 )
      wire#w1
      Coil( "CompALTA-MTA".FallaCompresor4 )
   END_RUNG
   RUNG wire#powerrail
      Contact( "DB_ALA_MEM".x88 )
   END_RUNG wire#w1
   RUNG wire#powerrail
      Contact( "DB_ALA_MEM".x89 )
   END_RUNG wire#w1
   RUNG wire#powerrail
      Contact( "DB_ALA_MEM".x90 )
   END_RUNG wire#w1
   RUNG wire#powerrail
      Contact( "DB_ALA_MEM".x74 )
   END_RUNG wire#w1
   RUNG wire#powerrail
      Contact( "DB_ALA_MEM".x75 )
   END_RUNG wire#w1
   RUNG wire#powerrail
      Contact( "DB_ALA_MEM".x133 )
   END_RUNG wire#w1
   RUNG wire#powerrail
      Contact( "FiltoPresostato_1".Q )
      Contact( "Enclavamientos".En1 )
      wire#w2
      I_Contact( "PanelCmpAlta".MantMC004 )
   END_RUNG wire#w1
   RUNG wire#powerrail
      Contact( "FallTempCritEnclav" )
      Contact( "Enclavamientos".En1 )
   END_RUNG wire#w2
   RUNG wire#powerrail
      Contact( "DB_ALA_PRE".x139 )
   END_RUNG wire#w1
   RUNG wire#w1
      R_Coil( "PanelCmpAlta".MarchaPanelMC004 )
   END_RUNG
   // the same network as SCL:
   "CompALTA-MTA".FallaCompresor4 := "DB_ALA_MEM".x87 OR "DB_ALA_MEM".x88 OR "DB_ALA_MEM".x89 OR "DB_ALA_MEM".x90 OR "DB_ALA_MEM".x74 OR "DB_ALA_MEM".x75 OR "DB_ALA_MEM".x133 OR ((("FiltoPresostato_1".Q AND "Enclavamientos".En1) OR ("FallTempCritEnclav" AND "Enclavamientos".En1)) AND NOT "PanelCmpAlta".MantMC004) OR "DB_ALA_PRE".x139;
   IF "CompALTA-MTA".FallaCompresor4 THEN "PanelCmpAlta".MarchaPanelMC004 := FALSE; END_IF;
END_REGION

REGION Network 9: Fallas de MC005 - Compresor de Alta ABC5
   RUNG wire#powerrail
      I_Contact( "PanelCmpAlta".MantMC005 )
      wire#w1
      Contact( "MC005_PTA" )
      Coil( "DB_ALA_PRE".x91 )
   END_RUNG
   RUNG wire#w1
      Contact( "MC005_PTB" )
      Coil( "DB_ALA_PRE".x92 )
   END_RUNG
   RUNG wire#w1
      Contact( "MC005_TTA" )
      Coil( "DB_ALA_PRE".x93 )
   END_RUNG
   RUNG wire#w1
      Contact( "MC005_TTB" )
      Coil( "DB_ALA_PRE".x94 )
   END_RUNG
   RUNG wire#w1
      Contact( "DB-PurgaComAlta".Habil_PurgaABC5 )
      Contact( "MC005_EVP" )
      I_Contact( "MC005_ConfPurga" )
      S_ODT(T_NO := "Tag_83", TV := S5Time#500ms, R :=, BI =>, RET_VAL =>)
      Coil( "DB_ALA_PRE".x140 )
   END_RUNG
   // the same network as SCL:
   #_w1 := NOT "PanelCmpAlta".MantMC005;
   "DB_ALA_PRE".x91 := #_w1 AND "MC005_PTA";
   "DB_ALA_PRE".x92 := #_w1 AND "MC005_PTB";
   "DB_ALA_PRE".x93 := #_w1 AND "MC005_TTA";
   "DB_ALA_PRE".x94 := #_w1 AND "MC005_TTB";
   #_s5time1 := S_ODT(T_NO := "Tag_83",
                      S := #_w1 AND "DB-PurgaComAlta".Habil_PurgaABC5 AND "MC005_EVP" AND NOT "MC005_ConfPurga",
                      TV := S5Time#500ms,
                      Q => #_w2);
   "DB_ALA_PRE".x140 := #_w2;
END_REGION

REGION Network 10: FallaCompresor5 (ABC5) / Alguna Falla en MC005 - Compresor de Alta ABC5